VERSION : 0.1
   VAR_TEMP
      Pump_A : Struct
         Cond_01 : Bool;   // Condition 01
         Cond_02 : Bool;
         Cond_03 : Bool;   // Condition 03
      END_STRUCT;
      Pump_B : Struct
         Cond_01 : Bool;   // Condition 01
         Cond_02 : Bool;   // Condition 02
         Cond_03 : Bool;   // Condition 03
      END_STRUCT;
   END_VAR
BEGIN
   //****** Equipmens Activation*******
   //
   //IF "AlwaysFALSE" THEN
       //**************************************************************
       //Feed Water Pump A
       // Condition to CmdOn "On Command" 
       IF "P-104A_DB".Config.HMI.Enable_HMI_Controls = 1 THEN
           #Pump_A.Cond_01 := "T-104_DB".Equipments."P-104A".Enable AND ("T-104_DB".PmpSel."P-104AB" = 1 OR "T-104_DB".PmpSel."P-104AB" = 3);
           #Pump_A.Cond_02 := "T-104_DB".ExchangeCmds.Receive.ReqWater; //Route Open to sent to the Reactor
           "T-104_DB".Equipments."P-104A".CmdOn := #Pump_A.Cond_01 AND #Pump_A.Cond_02 AND NOT "T-104_DB".Cmds.Hold;
           IF "T-104_DB".Equipments."P-104A".CmdOn THEN
               "P-104A_DB".Stop_CMD := False;
               "P-104A_DB".Start_CMD := true;
               "P-104A_DB".ON := TRUE;
               "P-104A_DB".OFF := FALSE;
           ELSE
               "P-104A_DB".Stop_CMD := true;
               "P-104A_DB".Start_CMD := false;
               "P-104A_DB".ON := FALSE;
               "P-104A_DB".OFF := TRUE;
           END_IF;
       END_IF;
       //**************************************************************
       //Feed Water Pump B
       // Condition to CmdOn "On Command" 
       IF "P-104B_DB".Config.HMI.Enable_HMI_Controls = 1 THEN
           #Pump_B.Cond_01 := "T-104_DB".Equipments."P-104B".Enable AND ("T-104_DB".PmpSel."P-104AB" = 2 OR "T-104_DB".PmpSel."P-104AB" = 3);
           #Pump_B.Cond_02 := "T-104_DB".ExchangeCmds.Receive.ReqWater; //Route Open to sent to the Reactor
           "T-104_DB".Equipments."P-104B".CmdOn := #Pump_B.Cond_01 AND #Pump_B.Cond_02 AND NOT "T-104_DB".Cmds.Hold AND "AlwaysFALSE";
           IF "T-104_DB".Equipments."P-104B".CmdOn THEN
               "P-104B_DB".ON := TRUE;
               "P-104B_DB".OFF := FALSE;
           ELSE
               "P-104B_DB".ON := FALSE;
               "P-104B_DB".OFF := TRUE;
           END_IF;
       END_IF;
   //END_IF;
   "T-104_DB".ExchangeCmds.Send.PumpingOut := ("P-104A_DB".CF AND ("PT-104A_DB".SAI>0.2)) OR ("P-104B_DB".CF AND ("PT-104B_DB".SAI>0.2));
   "T-104_DB".ExchangeCmds.Send.PumpsOff := NOT "P-104A_DB".CF AND NOT "P-104B_DB".CF;//AND ("PT-104A_DB".SAI<0.2)) AND (NOT "P-104B_DB".CF AND ("PT-104B_DB".SAI<0.2));
   //*****************************************Tank Ready********************************************************************
   "T-104_DB".ExchangeCmds.Send.TankReady := "T-104_DB".Status.Step = 21 AND "T-104_DB".PmpSel."P-104AB" > 0;
END_FUNCTION

FUNCTION "T-104_SignalsOutExchange" : Void   // FC87, LAD
{ S7_Optimized_Access := 'TRUE' }
VERSION : 0.1
BEGIN

REGION Network 1: Started (Send)
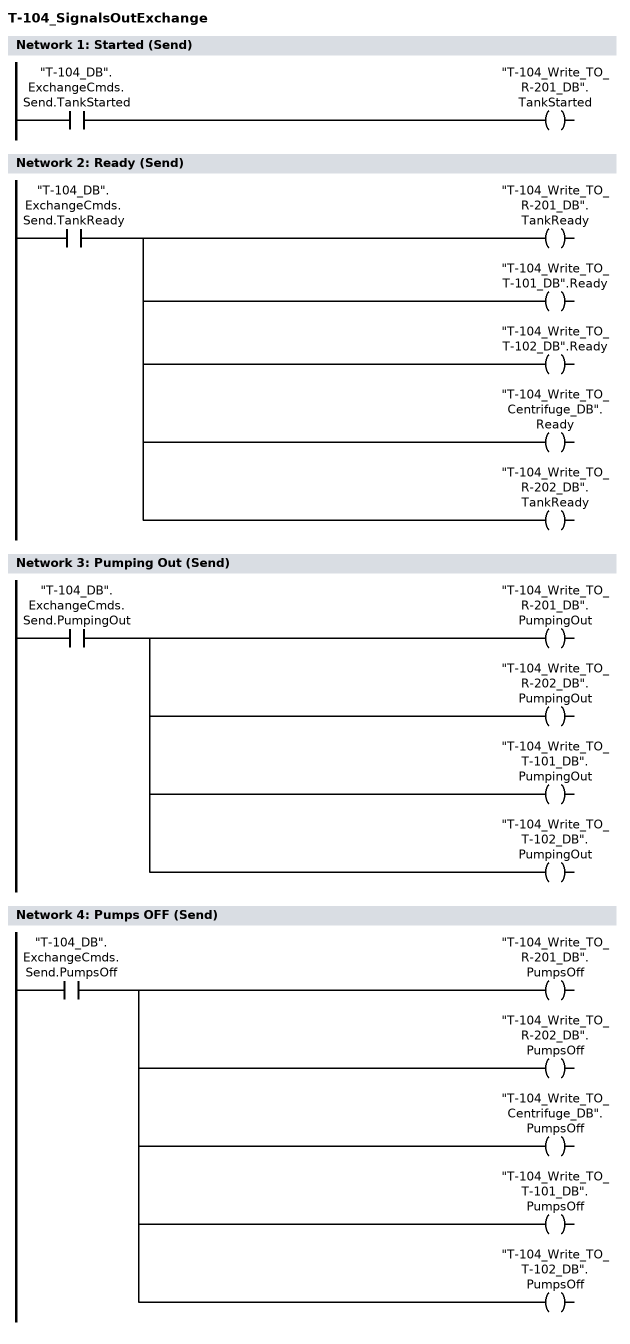
   RUNG wire#powerrail
      Contact( "T-104_DB".ExchangeCmds.Send.TankStarted )
      Coil( "T-104_Write_TO_R-201_DB".TankStarted )
   END_RUNG
   // the same network as SCL:
   "T-104_Write_TO_R-201_DB".TankStarted := "T-104_DB".ExchangeCmds.Send.TankStarted;
END_REGION

REGION Network 2: Ready (Send)
   RUNG wire#powerrail
      Contact( "T-104_DB".ExchangeCmds.Send.TankReady )
      wire#w1
      Coil( "T-104_Write_TO_R-201_DB".TankReady )
   END_RUNG
   RUNG wire#w1
      Coil( "T-104_Write_TO_T-101_DB".Ready )
   END_RUNG
   RUNG wire#w1
      Coil( "T-104_Write_TO_T-102_DB".Ready )
   END_RUNG
   RUNG wire#w1
      Coil( "T-104_Write_TO_Centrifuge_DB".Ready )
   END_RUNG
   RUNG wire#w1
      Coil( "T-104_Write_TO_R-202_DB".TankReady )
   END_RUNG
   // the same network as SCL:
   "T-104_Write_TO_R-201_DB".TankReady := "T-104_DB".ExchangeCmds.Send.TankReady;
   "T-104_Write_TO_T-101_DB".Ready := "T-104_DB".ExchangeCmds.Send.TankReady;
   "T-104_Write_TO_T-102_DB".Ready := "T-104_DB".ExchangeCmds.Send.TankReady;
   "T-104_Write_TO_Centrifuge_DB".Ready := "T-104_DB".ExchangeCmds.Send.TankReady;
   "T-104_Write_TO_R-202_DB".TankReady := "T-104_DB".ExchangeCmds.Send.TankReady;
END_REGION

REGION Network 3: Pumping Out (Send)
   RUNG wire#powerrail
      Contact( "T-104_DB".ExchangeCmds.Send.PumpingOut )
      wire#w1
      Coil( "T-104_Write_TO_R-201_DB".PumpingOut )
   END_RUNG
   RUNG wire#w1
      Coil( "T-104_Write_TO_R-202_DB".PumpingOut )
   END_RUNG
   RUNG wire#w1
      Coil( "T-104_Write_TO_T-101_DB".PumpingOut )
   END_RUNG
   RUNG wire#w1
      Coil( "T-104_Write_TO_T-102_DB".PumpingOut )
   END_RUNG
   // the same network as SCL:
   "T-104_Write_TO_R-201_DB".PumpingOut := "T-104_DB".ExchangeCmds.Send.PumpingOut;
   "T-104_Write_TO_R-202_DB".PumpingOut := "T-104_DB".ExchangeCmds.Send.PumpingOut;
   "T-104_Write_TO_T-101_DB".PumpingOut := "T-104_DB".ExchangeCmds.Send.PumpingOut;
   "T-104_Write_TO_T-102_DB".PumpingOut := "T-104_DB".ExchangeCmds.Send.PumpingOut;
END_REGION

REGION Network 4: Pumps OFF (Send)
   RUNG wire#powerrail
      Contact( "T-104_DB".ExchangeCmds.Send.PumpsOff )
      wire#w1
      Coil( "T-104_Write_TO_R-201_DB".PumpsOff )
   END_RUNG
   RUNG wire#w1
      Coil( "T-104_Write_TO_R-202_DB".PumpsOff )
   END_RUNG
   RUNG wire#w1
      Coil( "T-104_Write_TO_Centrifuge_DB".PumpsOff )
   END_RUNG
   RUNG wire#w1
      Coil( "T-104_Write_TO_T-101_DB".PumpsOff )
   END_RUNG
   RUNG wire#w1
      Coil( "T-104_Write_TO_T-102_DB".PumpsOff )
   END_RUNG
   // the same network as SCL:
   "T-104_Write_TO_R-201_DB".PumpsOff := "T-104_DB".ExchangeCmds.Send.PumpsOff;
   "T-104_Write_TO_R-202_DB".PumpsOff := "T-104_DB".ExchangeCmds.Send.PumpsOff;
   "T-104_Write_TO_Centrifuge_DB".PumpsOff := "T-104_DB".ExchangeCmds.Send.PumpsOff;
   "T-104_Write_TO_T-101_DB".PumpsOff := "T-104_DB".ExchangeCmds.Send.PumpsOff;
   "T-104_Write_TO_T-102_DB".PumpsOff := "T-104_DB".ExchangeCmds.Send.PumpsOff;
END_REGION
END_FUNCTION

FUNCTION "T-104_SEQ_FC" : Void   // FC88, LAD
{ S7_Optimized_Access := 'TRUE' }
VERSION : 0.1
   VAR_TEMP   // added for the SCL form of the ladder/FBD networks
      _w1 : Bool;
   END_VAR
BEGIN

REGION Network 2: Abort
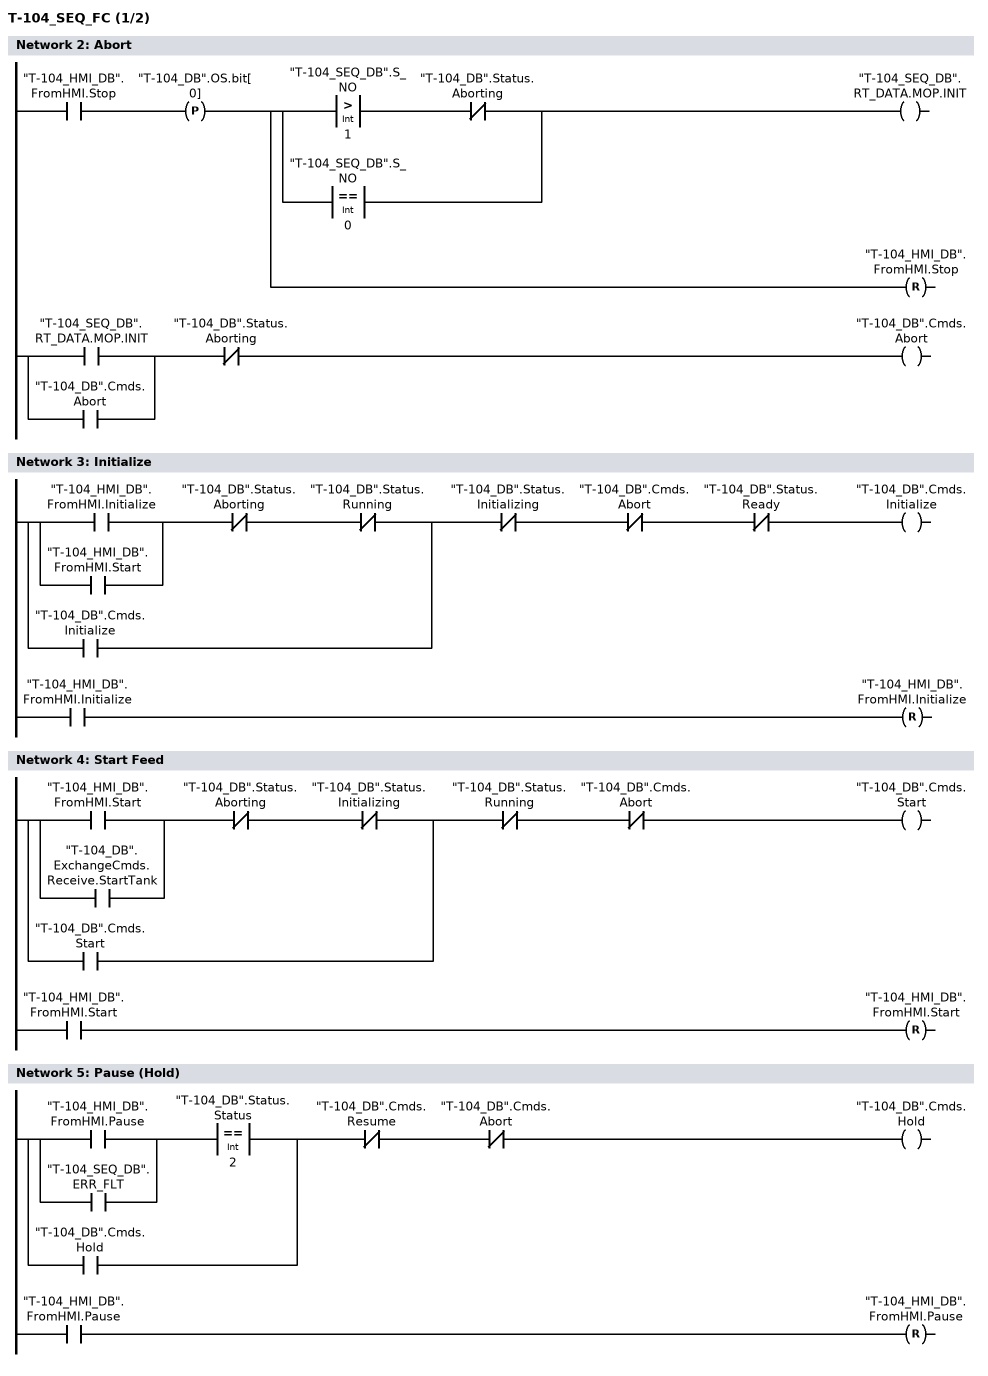
   RUNG wire#powerrail
      Contact( "T-104_HMI_DB".FromHMI.Stop )
      P_Trig( "T-104_DB".OS.bit[0] )
      wire#w1
      { S7_Templates := "SrcType := Int" } GT_Contact(in1 := "T-104_SEQ_DB".S_NO, in2 := 1)
      I_Contact( "T-104_DB".Status.Aborting )
      wire#w2
      Coil( "T-104_SEQ_DB".RT_DATA.MOP.INIT )
   END_RUNG
   RUNG wire#w1
      { S7_Templates := "SrcType := Int" } EQ_Contact(in1 := "T-104_SEQ_DB".S_NO, in2 := 0)
   END_RUNG wire#w2
   RUNG wire#w1
      R_Coil( "T-104_HMI_DB".FromHMI.Stop )
   END_RUNG
   RUNG wire#powerrail
      Contact( "T-104_SEQ_DB".RT_DATA.MOP.INIT )
      wire#w3
      I_Contact( "T-104_DB".Status.Aborting )
      Coil( "T-104_DB".Cmds.Abort )
   END_RUNG
   RUNG wire#powerrail
      Contact( "T-104_DB".Cmds.Abort )
   END_RUNG wire#w3
   // the same network as SCL:
   #_w1 := "T-104_HMI_DB".FromHMI.Stop AND NOT "T-104_DB".OS.bit[0];   // rising edge
   "T-104_DB".OS.bit[0] := "T-104_HMI_DB".FromHMI.Stop;
   "T-104_SEQ_DB".RT_DATA.MOP.INIT := #_w1 AND ((("T-104_SEQ_DB".S_NO > 1) AND NOT "T-104_DB".Status.Aborting) OR ("T-104_SEQ_DB".S_NO = 0));
   IF #_w1 THEN "T-104_HMI_DB".FromHMI.Stop := FALSE; END_IF;
   "T-104_DB".Cmds.Abort := ("T-104_SEQ_DB".RT_DATA.MOP.INIT OR "T-104_DB".Cmds.Abort) AND NOT "T-104_DB".Status.Aborting;
END_REGION

REGION Network 3: Initialize
   RUNG wire#powerrail
      Contact( "T-104_HMI_DB".FromHMI.Initialize )
      wire#w1
      I_Contact( "T-104_DB".Status.Aborting )
      I_Contact( "T-104_DB".Status.Running )
      wire#w2
      I_Contact( "T-104_DB".Status.Initializing )
      I_Contact( "T-104_DB".Cmds.Abort )
      I_Contact( "T-104_DB".Status.Ready )
      Coil( "T-104_DB".Cmds.Initialize )
   END_RUNG
   RUNG wire#powerrail
      Contact( "T-104_HMI_DB".FromHMI.Start )
   END_RUNG wire#w1
   RUNG wire#powerrail
      Contact( "T-104_DB".Cmds.Initialize )
   END_RUNG wire#w2
   RUNG wire#powerrail
      Contact( "T-104_HMI_DB".FromHMI.Initialize )
      R_Coil( "T-104_HMI_DB".FromHMI.Initialize )
   END_RUNG
   // the same network as SCL:
   "T-104_DB".Cmds.Initialize := ((("T-104_HMI_DB".FromHMI.Initialize OR "T-104_HMI_DB".FromHMI.Start) AND NOT "T-104_DB".Status.Aborting AND NOT "T-104_DB".Status.Running) OR "T-104_DB".Cmds.Initialize) AND NOT "T-104_DB".Status.Initializing AND NOT "T-104_DB".Cmds.Abort AND NOT "T-104_DB".Status.Ready;
   IF "T-104_HMI_DB".FromHMI.Initialize THEN "T-104_HMI_DB".FromHMI.Initialize := FALSE; END_IF;
END_REGION

REGION Network 4: Start Feed
   RUNG wire#powerrail
      Contact( "T-104_HMI_DB".FromHMI.Start )
      wire#w1
      I_Contact( "T-104_DB".Status.Aborting )
      I_Contact( "T-104_DB".Status.Initializing )
      wire#w2
      I_Contact( "T-104_DB".Status.Running )
      I_Contact( "T-104_DB".Cmds.Abort )
      Coil( "T-104_DB".Cmds.Start )
   END_RUNG
   RUNG wire#powerrail
      Contact( "T-104_DB".ExchangeCmds.Receive.StartTank )
   END_RUNG wire#w1
   RUNG wire#powerrail
      Contact( "T-104_DB".Cmds.Start )
   END_RUNG wire#w2
   RUNG wire#powerrail
      Contact( "T-104_HMI_DB".FromHMI.Start )
      R_Coil( "T-104_HMI_DB".FromHMI.Start )
   END_RUNG
   // the same network as SCL:
   "T-104_DB".Cmds.Start := ((("T-104_HMI_DB".FromHMI.Start OR "T-104_DB".ExchangeCmds.Receive.StartTank) AND NOT "T-104_DB".Status.Aborting AND NOT "T-104_DB".Status.Initializing) OR "T-104_DB".Cmds.Start) AND NOT "T-104_DB".Status.Running AND NOT "T-104_DB".Cmds.Abort;
   IF "T-104_HMI_DB".FromHMI.Start THEN "T-104_HMI_DB".FromHMI.Start := FALSE; END_IF;
END_REGION

REGION Network 5: Pause (Hold)
   RUNG wire#powerrail
      Contact( "T-104_HMI_DB".FromHMI.Pause )
      wire#w1
      { S7_Templates := "SrcType := Int" } EQ_Contact(in1 := "T-104_DB".Status.Status, in2 := 2)
      wire#w2
      I_Contact( "T-104_DB".Cmds.Resume )
      I_Contact( "T-104_DB".Cmds.Abort )
      Coil( "T-104_DB".Cmds.Hold )
   END_RUNG
   RUNG wire#powerrail
      Contact( "T-104_SEQ_DB".ERR_FLT )
   END_RUNG wire#w1
   RUNG wire#powerrail
      Contact( "T-104_DB".Cmds.Hold )
   END_RUNG wire#w2
   RUNG wire#powerrail
      Contact( "T-104_HMI_DB".FromHMI.Pause )
      R_Coil( "T-104_HMI_DB".FromHMI.Pause )
   END_RUNG
   // the same network as SCL:
   "T-104_DB".Cmds.Hold := ((("T-104_HMI_DB".FromHMI.Pause OR "T-104_SEQ_DB".ERR_FLT) AND ("T-104_DB".Status.Status = 2)) OR "T-104_DB".Cmds.Hold) AND NOT "T-104_DB".Cmds.Resume AND NOT "T-104_DB".Cmds.Abort;
   IF "T-104_HMI_DB".FromHMI.Pause THEN "T-104_HMI_DB".FromHMI.Pause := FALSE; END_IF;
END_REGION

REGION Network 6: Restart From Pause (Hold)
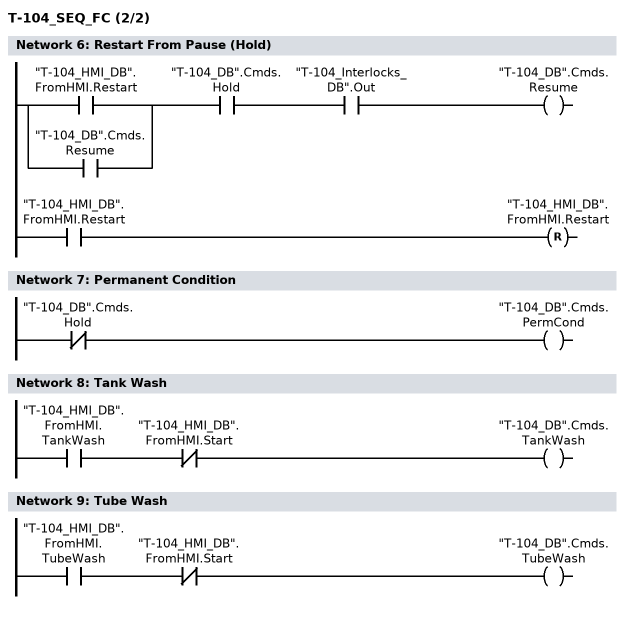
   RUNG wire#powerrail
      Contact( "T-104_HMI_DB".FromHMI.Restart )
      wire#w1
      Contact( "T-104_DB".Cmds.Hold )
      Contact( "T-104_Interlocks_DB".Out )
      Coil( "T-104_DB".Cmds.Resume )
   END_RUNG
   RUNG wire#powerrail
      Contact( "T-104_DB".Cmds.Resume )
   END_RUNG wire#w1
   RUNG wire#powerrail
      Contact( "T-104_HMI_DB".FromHMI.Restart )
      R_Coil( "T-104_HMI_DB".FromHMI.Restart )
   END_RUNG
   // the same network as SCL:
   "T-104_DB".Cmds.Resume := ("T-104_HMI_DB".FromHMI.Restart OR "T-104_DB".Cmds.Resume) AND "T-104_DB".Cmds.Hold AND "T-104_Interlocks_DB".Out;
   IF "T-104_HMI_DB".FromHMI.Restart THEN "T-104_HMI_DB".FromHMI.Restart := FALSE; END_IF;
END_REGION

REGION Network 7: Permanent Condition
   RUNG wire#powerrail
      I_Contact( "T-104_DB".Cmds.Hold )
      Coil( "T-104_DB".Cmds.PermCond )
   END_RUNG
   // the same network as SCL:
   "T-104_DB".Cmds.PermCond := NOT "T-104_DB".Cmds.Hold;
END_REGION

REGION Network 8: Tank Wash
   RUNG wire#powerrail
      Contact( "T-104_HMI_DB".FromHMI.TankWash )
      I_Contact( "T-104_HMI_DB".FromHMI.Start )
      Coil( "T-104_DB".Cmds.TankWash )
   END_RUNG
   // the same network as SCL:
   "T-104_DB".Cmds.TankWash := "T-104_HMI_DB".FromHMI.TankWash AND NOT "T-104_HMI_DB".FromHMI.Start;
END_REGION

REGION Network 9: Tube Wash
   RUNG wire#powerrail
      Contact( "T-104_HMI_DB".FromHMI.TubeWash )
      I_Contact( "T-104_HMI_DB".FromHMI.Start )
      Coil( "T-104_DB".Cmds.TubeWash )
   END_RUNG
   // the same network as SCL:
   "T-104_DB".Cmds.TubeWash := "T-104_HMI_DB".FromHMI.TubeWash AND NOT "T-104_HMI_DB".FromHMI.Start;
END_REGION

REGION Network 10 (SCL): Sequence Status
   IF "T-104_SEQ_DB".S_NO= 1 THEN
       "T-104_DB".Status.Status := 1; //Idle
   ELSIF "T-104_SEQ_DB".S_NO > 1 AND "T-104_SEQ_DB".S_NO < 150 AND NOT "T-104_SEQ_DB".ERR_FLT AND NOT "T-104_DB".Cmds.Hold THEN
       "T-104_DB".Status.Status := 2; //Running
   ELSIF "T-104_SEQ_DB".S_NO >= 151 AND "T-104_SEQ_DB".S_NO <= 160 AND NOT "T-104_SEQ_DB".ERR_FLT THEN
       "T-104_DB".Status.Status := 3; // Stopping
   ELSIF  "T-104_SEQ_DB".ERR_FLT AND  ("T-104_SEQ_DB".S_NO > 1 AND "T-104_SEQ_DB".S_NO < 150) THEN
       "T-104_DB".Status.Status := 4; // Held
   ELSIF  "T-104_SEQ_DB".ERR_FLT AND  ("T-104_SEQ_DB".S_NO > 1 AND "T-104_SEQ_DB".S_NO < 150) AND "T-104_Aux_DB"."Bool".TOff  THEN
       "T-104_DB".Status.Status := 5; // Holding
   ELSE
       "T-104_DB".Status.Status := 6; // Unknown
   END_IF;

   "T-104_DB".Status.Running := ("T-104_SEQ_DB".S_NO > 3 AND "T-104_SEQ_DB".S_NO <= 150);
   "T-104_DB".Status.Initializing := ("T-104_SEQ_DB".S_NO >= 141 AND "T-104_SEQ_DB".S_NO <= 150);

   //Enable/Disable HMI Start/Stop Button
   "T-104_HMI_DB".ToHMI.EnStopButton := ("T-104_DB".Status.Status > 1) OR "T-104_DB".Status.Step = 0; //Enable HMI Stop Button
   "T-104_HMI_DB".ToHMI.EnStartButton := "T-104_DB".Status.Status = 1; //Idle
   "T-104_HMI_DB".ToHMI.EnPauseButton := "T-104_DB".Status.Status = 2; //Enable Pause Button
   "T-104_HMI_DB".ToHMI.EnRestartButton :=  "T-104_DB".Status.Status = 4; //Enable Restart Button

   //****Interlock Activated
   "T-104_HMI_DB".ToHMI.InterlockActivated := "T-104_Interlocks_DB".Out;
END_REGION

REGION Network 11 (SCL): Sequence Step
   "T-104_DB".Status.Step := "T-104_SEQ_DB".S_NO;
END_REGION

REGION Network 12 (SCL): Sequence state (Procedure running)
   IF "T-104_SEQ_DB".S_NO = 3 OR "T-104_SEQ_DB".S_NO = 4 THEN
       "T-104_DB".Status.State := 1; //Ready
   ELSIF "T-104_SEQ_DB".S_NO >= 21 AND "T-104_SEQ_DB".S_NO <= 60 THEN
       "T-104_DB".Status.State := 2; //Mixing 
   ELSIF "T-104_SEQ_DB".S_NO >= 61 AND "T-104_SEQ_DB".S_NO <= 80 THEN
       "T-104_DB".Status.State := 3; //Pouring
   ELSIF "T-104_SEQ_DB".S_NO >= 141 AND "T-104_SEQ_DB".S_NO <= 150 THEN
       "T-104_DB".Status.State := 4; //Initializing
   ELSIF "T-104_SEQ_DB".S_NO >= 151 AND "T-104_SEQ_DB".S_NO <= 160 THEN
       "T-104_DB".Status.State := 5; //Aborting
   ELSE
       "T-104_DB".Status.State := 0;
   END_IF;
END_REGION

REGION Network 13: Sequence State
END_REGION
END_FUNCTION

// folder: State MACHINE/1)Tanks/Tank T-104 (Water System)/T-104 <---> Centrifuge

FUNCTION "T-104_Signals_FROM_Centrifuge" : Void   // FC71, LAD
{ S7_Optimized_Access := 'TRUE' }
VERSION : 0.1
BEGIN

REGION Network 1: Start Sequence
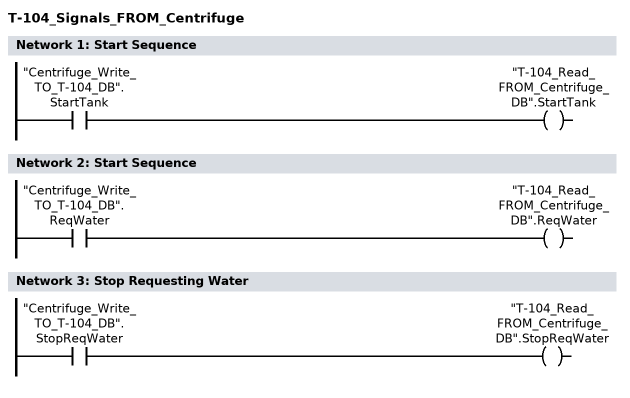
   RUNG wire#powerrail
      Contact( "Centrifuge_Write_TO_T-104_DB".StartTank )
      Coil( "T-104_Read_FROM_Centrifuge_DB".StartTank )
   END_RUNG
   // the same network as SCL:
   "T-104_Read_FROM_Centrifuge_DB".StartTank := "Centrifuge_Write_TO_T-104_DB".StartTank;
END_REGION

REGION Network 2: Start Sequence
   RUNG wire#powerrail
      Contact( "Centrifuge_Write_TO_T-104_DB".ReqWater )
      Coil( "T-104_Read_FROM_Centrifuge_DB".ReqWater )
   END_RUNG
   // the same network as SCL:
   "T-104_Read_FROM_Centrifuge_DB".ReqWater := "Centrifuge_Write_TO_T-104_DB".ReqWater;
END_REGION

REGION Network 3: Stop Requesting Water
   RUNG wire#powerrail
      Contact( "Centrifuge_Write_TO_T-104_DB".StopReqWater )
      Coil( "T-104_Read_FROM_Centrifuge_DB".StopReqWater )
   END_RUNG
   // the same network as SCL:
   "T-104_Read_FROM_Centrifuge_DB".StopReqWater := "Centrifuge_Write_TO_T-104_DB".StopReqWater;
END_REGION
END_FUNCTION

// folder: State MACHINE/1)Tanks/Tank T-104 (Water System)/T-104 <---> R-201

FUNCTION "T-104_Signals_FROM_R-201" : Void   // FC50, LAD
{ S7_Optimized_Access := 'TRUE' }
VERSION : 0.1
BEGIN

REGION Network 1: Start Sequence
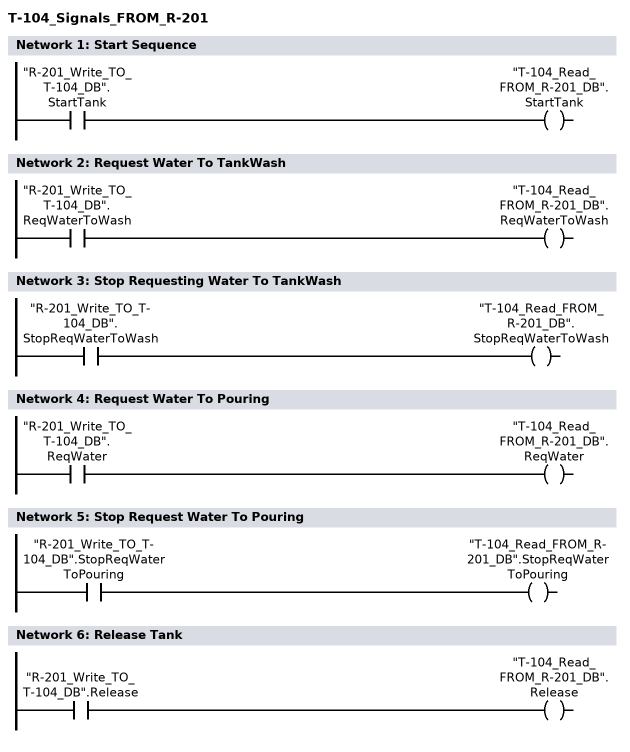
   RUNG wire#powerrail
      Contact( "R-201_Write_TO_T-104_DB".StartTank )
      Coil( "T-104_Read_FROM_R-201_DB".StartTank )
   END_RUNG
   // the same network as SCL:
   "T-104_Read_FROM_R-201_DB".StartTank := "R-201_Write_TO_T-104_DB".StartTank;
END_REGION

REGION Network 2: Request Water To TankWash
   RUNG wire#powerrail
      Contact( "R-201_Write_TO_T-104_DB".ReqWaterToWash )
      Coil( "T-104_Read_FROM_R-201_DB".ReqWaterToWash )
   END_RUNG
   // the same network as SCL:
   "T-104_Read_FROM_R-201_DB".ReqWaterToWash := "R-201_Write_TO_T-104_DB".ReqWaterToWash;
END_REGION

REGION Network 3: Stop Requesting Water To TankWash
   RUNG wire#powerrail
      Contact( "R-201_Write_TO_T-104_DB".StopReqWaterToWash )
      Coil( "T-104_Read_FROM_R-201_DB".StopReqWaterToWash )
   END_RUNG
   // the same network as SCL:
   "T-104_Read_FROM_R-201_DB".StopReqWaterToWash := "R-201_Write_TO_T-104_DB".StopReqWaterToWash;
END_REGION

REGION Network 4: Request Water To Pouring
   RUNG wire#powerrail
      Contact( "R-201_Write_TO_T-104_DB".ReqWater )
      Coil( "T-104_Read_FROM_R-201_DB".ReqWater )
   END_RUNG
   // the same network as SCL:
   "T-104_Read_FROM_R-201_DB".ReqWater := "R-201_Write_TO_T-104_DB".ReqWater;
END_REGION

REGION Network 5: Stop Request Water To Pouring
   RUNG wire#powerrail
      Contact( "R-201_Write_TO_T-104_DB".StopReqWaterToPouring )
      Coil( "T-104_Read_FROM_R-201_DB".StopReqWaterToPouring )
   END_RUNG
   // the same network as SCL:
   "T-104_Read_FROM_R-201_DB".StopReqWaterToPouring := "R-201_Write_TO_T-104_DB".StopReqWaterToPouring;
END_REGION

REGION Network 6: Release Tank
   RUNG wire#powerrail
      Contact( "R-201_Write_TO_T-104_DB".Release )
      Coil( "T-104_Read_FROM_R-201_DB".Release )
   END_RUNG
   // the same network as SCL:
   "T-104_Read_FROM_R-201_DB".Release := "R-201_Write_TO_T-104_DB".Release;
END_REGION
END_FUNCTION

// folder: State MACHINE/1)Tanks/Tank T-104 (Water System)/T-104 <---> R-202

FUNCTION "T-104_Signals_FROM_R-202" : Void   // FC72, LAD
{ S7_Optimized_Access := 'TRUE' }
VERSION : 0.1
BEGIN

REGION Network 1: Start Sequence
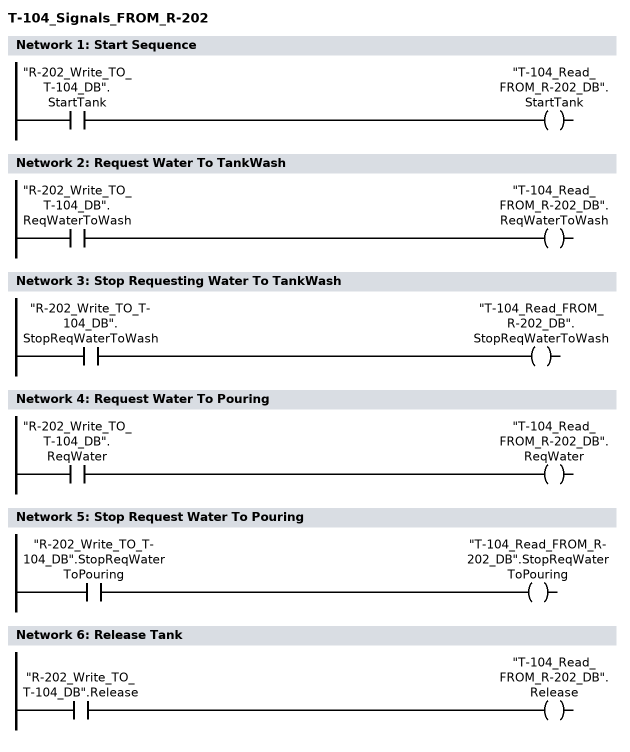
   RUNG wire#powerrail
      Contact( "R-202_Write_TO_T-104_DB".StartTank )
      Coil( "T-104_Read_FROM_R-202_DB".StartTank )
   END_RUNG
   // the same network as SCL:
   "T-104_Read_FROM_R-202_DB".StartTank := "R-202_Write_TO_T-104_DB".StartTank;
END_REGION

REGION Network 2: Request Water To TankWash
   RUNG wire#powerrail
      Contact( "R-202_Write_TO_T-104_DB".ReqWaterToWash )
      Coil( "T-104_Read_FROM_R-202_DB".ReqWaterToWash )
   END_RUNG
   // the same network as SCL:
   "T-104_Read_FROM_R-202_DB".ReqWaterToWash := "R-202_Write_TO_T-104_DB".ReqWaterToWash;
END_REGION

REGION Network 3: Stop Requesting Water To TankWash
   RUNG wire#powerrail
      Contact( "R-202_Write_TO_T-104_DB".StopReqWaterToWash )
      Coil( "T-104_Read_FROM_R-202_DB".StopReqWaterToWash )
   END_RUNG
   // the same network as SCL:
   "T-104_Read_FROM_R-202_DB".StopReqWaterToWash := "R-202_Write_TO_T-104_DB".StopReqWaterToWash;
END_REGION

REGION Network 4: Request Water To Pouring
   RUNG wire#powerrail
      Contact( "R-202_Write_TO_T-104_DB".ReqWater )
      Coil( "T-104_Read_FROM_R-202_DB".ReqWater )
   END_RUNG
   // the same network as SCL:
   "T-104_Read_FROM_R-202_DB".ReqWater := "R-202_Write_TO_T-104_DB".ReqWater;
END_REGION

REGION Network 5: Stop Request Water To Pouring
   RUNG wire#powerrail
      Contact( "R-202_Write_TO_T-104_DB".StopReqWaterToPouring )
      Coil( "T-104_Read_FROM_R-202_DB".StopReqWaterToPouring )
   END_RUNG
   // the same network as SCL:
   "T-104_Read_FROM_R-202_DB".StopReqWaterToPouring := "R-202_Write_TO_T-104_DB".StopReqWaterToPouring;
END_REGION

REGION Network 6: Release Tank
   RUNG wire#powerrail
      Contact( "R-202_Write_TO_T-104_DB".Release )
      Coil( "T-104_Read_FROM_R-202_DB".Release )
   END_RUNG
   // the same network as SCL:
   "T-104_Read_FROM_R-202_DB".Release := "R-202_Write_TO_T-104_DB".Release;
END_REGION
END_FUNCTION

// folder: State MACHINE/1)Tanks/Tank T-104 (Water System)/T-104 <---> T-101

FUNCTION "T-104_Signals_FROM_T-101" : Void   // FC74, LAD
{ S7_Optimized_Access := 'TRUE' }
VERSION : 0.1
BEGIN

REGION Network 1: Start Sequence
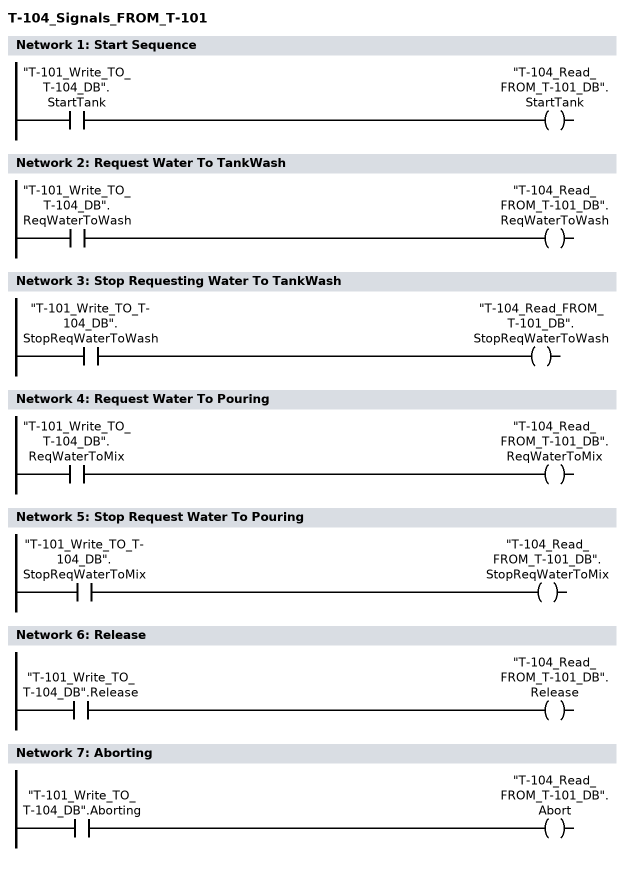
   RUNG wire#powerrail
      Contact( "T-101_Write_TO_T-104_DB".StartTank )
      Coil( "T-104_Read_FROM_T-101_DB".StartTank )
   END_RUNG
   // the same network as SCL:
   "T-104_Read_FROM_T-101_DB".StartTank := "T-101_Write_TO_T-104_DB".StartTank;
END_REGION

REGION Network 2: Request Water To TankWash
   RUNG wire#powerrail
      Contact( "T-101_Write_TO_T-104_DB".ReqWaterToWash )
      Coil( "T-104_Read_FROM_T-101_DB".ReqWaterToWash )
   END_RUNG
   // the same network as SCL:
   "T-104_Read_FROM_T-101_DB".ReqWaterToWash := "T-101_Write_TO_T-104_DB".ReqWaterToWash;
END_REGION

REGION Network 3: Stop Requesting Water To TankWash
   RUNG wire#powerrail
      Contact( "T-101_Write_TO_T-104_DB".StopReqWaterToWash )
      Coil( "T-104_Read_FROM_T-101_DB".StopReqWaterToWash )
   END_RUNG
   // the same network as SCL:
   "T-104_Read_FROM_T-101_DB".StopReqWaterToWash := "T-101_Write_TO_T-104_DB".StopReqWaterToWash;
END_REGION

REGION Network 4: Request Water To Pouring
   RUNG wire#powerrail
      Contact( "T-101_Write_TO_T-104_DB".ReqWaterToMix )
      Coil( "T-104_Read_FROM_T-101_DB".ReqWaterToMix )
   END_RUNG
   // the same network as SCL:
   "T-104_Read_FROM_T-101_DB".ReqWaterToMix := "T-101_Write_TO_T-104_DB".ReqWaterToMix;
END_REGION

REGION Network 5: Stop Request Water To Pouring
   RUNG wire#powerrail
      Contact( "T-101_Write_TO_T-104_DB".StopReqWaterToMix )
      Coil( "T-104_Read_FROM_T-101_DB".StopReqWaterToMix )
   END_RUNG
   // the same network as SCL:
   "T-104_Read_FROM_T-101_DB".StopReqWaterToMix := "T-101_Write_TO_T-104_DB".StopReqWaterToMix;
END_REGION

REGION Network 6: Release
   RUNG wire#powerrail
      Contact( "T-101_Write_TO_T-104_DB".Release )
      Coil( "T-104_Read_FROM_T-101_DB".Release )
   END_RUNG
   // the same network as SCL:
   "T-104_Read_FROM_T-101_DB".Release := "T-101_Write_TO_T-104_DB".Release;
END_REGION

REGION Network 7: Aborting
   RUNG wire#powerrail
      Contact( "T-101_Write_TO_T-104_DB".Aborting )
      Coil( "T-104_Read_FROM_T-101_DB".Abort )
   END_RUNG
   // the same network as SCL:
   "T-104_Read_FROM_T-101_DB".Abort := "T-101_Write_TO_T-104_DB".Aborting;
END_REGION
END_FUNCTION

// folder: State MACHINE/1)Tanks/Tank T-104 (Water System)/T-104 <---> T-102

FUNCTION "T-104_Signals_FROM_T-102" : Void   // FC73, LAD
{ S7_Optimized_Access := 'TRUE' }
VERSION : 0.1
BEGIN

REGION Network 1: Start Sequence
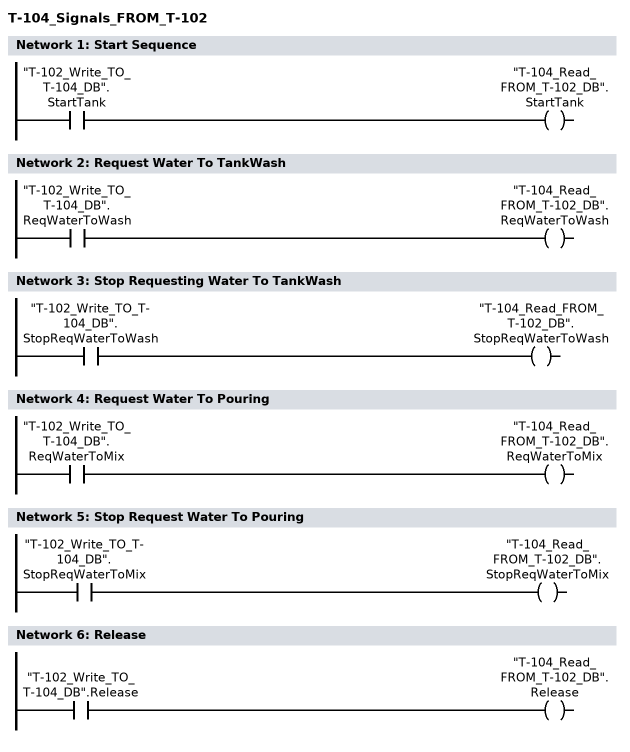
   RUNG wire#powerrail
      Contact( "T-102_Write_TO_T-104_DB".StartTank )
      Coil( "T-104_Read_FROM_T-102_DB".StartTank )
   END_RUNG
   // the same network as SCL:
   "T-104_Read_FROM_T-102_DB".StartTank := "T-102_Write_TO_T-104_DB".StartTank;
END_REGION

REGION Network 2: Request Water To TankWash
   RUNG wire#powerrail
      Contact( "T-102_Write_TO_T-104_DB".ReqWaterToWash )
      Coil( "T-104_Read_FROM_T-102_DB".ReqWaterToWash )
   END_RUNG
   // the same network as SCL:
   "T-104_Read_FROM_T-102_DB".ReqWaterToWash := "T-102_Write_TO_T-104_DB".ReqWaterToWash;
END_REGION

REGION Network 3: Stop Requesting Water To TankWash
   RUNG wire#powerrail
      Contact( "T-102_Write_TO_T-104_DB".StopReqWaterToWash )
      Coil( "T-104_Read_FROM_T-102_DB".StopReqWaterToWash )
   END_RUNG
   // the same network as SCL:
   "T-104_Read_FROM_T-102_DB".StopReqWaterToWash := "T-102_Write_TO_T-104_DB".StopReqWaterToWash;
END_REGION

REGION Network 4: Request Water To Pouring
   RUNG wire#powerrail
      Contact( "T-102_Write_TO_T-104_DB".ReqWaterToMix )
      Coil( "T-104_Read_FROM_T-102_DB".ReqWaterToMix )
   END_RUNG
   // the same network as SCL:
   "T-104_Read_FROM_T-102_DB".ReqWaterToMix := "T-102_Write_TO_T-104_DB".ReqWaterToMix;
END_REGION

REGION Network 5: Stop Request Water To Pouring
   RUNG wire#powerrail
      Contact( "T-102_Write_TO_T-104_DB".StopReqWaterToMix )
      Coil( "T-104_Read_FROM_T-102_DB".StopReqWaterToMix )
   END_RUNG
   // the same network as SCL:
   "T-104_Read_FROM_T-102_DB".StopReqWaterToMix := "T-102_Write_TO_T-104_DB".StopReqWaterToMix;
END_REGION

REGION Network 6: Release
   RUNG wire#powerrail
      Contact( "T-102_Write_TO_T-104_DB".Release )
      Coil( "T-104_Read_FROM_T-102_DB".Release )
   END_RUNG
   // the same network as SCL:
   "T-104_Read_FROM_T-102_DB".Release := "T-102_Write_TO_T-104_DB".Release;
END_REGION
END_FUNCTION

// folder: State MACHINE/2)Reactors/Reactor R-201

FUNCTION_BLOCK "R-201_SEQ"   // FB32, GRAPH_PLUS
{ S7_Optimized_Access := 'TRUE' }
VERSION : 0.1
   VAR_INPUT
      OFF_SQ : Bool := false;   // Turn sequence off
      INIT_SQ : Bool := false;   // Set sequence to initial state
      ACK_EF : Bool := false;   // Acknowledge all errors and faults
   END_VAR
   VAR_OUTPUT
      S_NO : Int := 0;   // Step number
      S_MORE : Bool := false;   // More steps are available and can be shown in S_NO
      S_ACTIVE : Bool := false;   // Step indicated in S_NO is active
      ERR_FLT : Bool := false;   // Interlock or supervision group error
      AUTO_ON : Bool := false;   // Automatic mode is active
   END_VAR
   VAR
      Reactor : Struct   // Reactor Ctrl
         IDLE : Bool;
         INITIALIZATION : Bool;   // Sequence initialization
         START : Bool;
         DONE_REACTING : Bool;
         COMPLETE : Bool;   // Reactor Complete Read only
         PARA : Bool;   // PARA load Batch side button
         ABORTING : Bool;   // Sequence about
         WAIT : Bool;   // Wating for Permissive read only
      END_STRUCT;
      "Aux Reactor" : Struct
         INITIALIZATION : Bool;
         START : Bool;
         DONE : Bool;
         COMPLETE : Bool;
         PARA : Bool;
         "SELECT_R-201" : Bool;
         "SELECT_R-202" : Bool;
         "SELECT_R-201/R-202" : Bool;
         "SELECT_R-201_T-103" : Bool;
         "SELECT_R-202_T-103" : Bool;
         ABORT : Bool;
         WAIT : Bool;
         LV : Bool;
         FLOW : Bool;
         MIX : Bool;
         "Pre-MIX" : Bool;
         REACTOR : Bool;
         WASH : Bool;
         TUBE : Bool;
         "SEQ_R-201" : Bool;
         "SEQ_R-202" : Bool;
         "SEQ_ R-201 & R-202" : Bool;
         "SEQ_T-103_R-201" : Bool;
         "SEQ_T-103_R-202" : Bool;
         BatchVolume : Real;
         Batchsize : Real;
         batchFlow : Real := 1.0;
         "batchFlow_T-102" : Real;
         BatchPH : Real := 7.0;
         "T-101" : Real;
         BatchTemp : Real := 80.0;
         PM : Bool;
         "TIME" : Struct
            "PRE-MIX" : Time;
            PH_DELAY : Time;
            REACTOR : Time;
            WATCH : Time;
            TUBE : Time;
            CountDown : Struct
               "PRE-MIX" : Time;
               PH_DELAY : Time;
               REACTOR : Time;
               WATCH : Time;
               TUBE : Time;
            END_STRUCT;
         END_STRUCT;
         "TIMER" : Struct
            "PRE-MIX" : IEC_TIMER;
            MIX : IEC_TIMER;
            PH_DELAY : IEC_TIMER;
            REACTOR : IEC_TIMER;
            WASH : IEC_TIMER;
            TUBE : IEC_TIMER;
         END_STRUCT;
      END_STRUCT;
      TEMP : Struct
         TANKS_BATCH : Real;
         "EMPTY_LV_0%" : Real;
         "MIN_LV_20%" : Real;
         "MAX_LV_80%" : Real;
         "BELOW_32%" : Real;
         "Greater_8%" : Real;
         "PRE-ADD" : Real;
         X_SOL_SIZE : Real;
         Y_SOL_SIZE : Real;
         PH_MIN : Real;
         PH_MAX : Real;
         OFFSEt : Struct
            MAX : Real;
            MIN : Real;
         END_STRUCT;
      END_STRUCT;
      COOLING : Struct   // Reactor Ctrl
         IDLE : Bool;
      END_STRUCT;
      HMI_INFO : Array[0..16] of UInt;
      IF_PAR : G7_IfParPlus_V6;
      RT_DATA : G7_RTDataPlus_V6;   // Internal data area
      Abort : G7_TransitionPlus_V6;   // Transition structure
      InitializeR : G7_TransitionPlus_V6;   // Transition structure
      "Fill/Pouring" : G7_TransitionPlus_V6;   // Transition structure
      Re : G7_TransitionPlus_V6;   // Transition structure
      "Fill/Pour" : G7_TransitionPlus_V6;   // Transition structure
      WashT : G7_TransitionPlus_V6;   // Transition structure
      WashTub : G7_TransitionPlus_V6;   // Transition structure
      Std : G7_TransitionPlus_V6;   // Transition structure
      StT : G7_TransitionPlus_V6;   // Transition structure
      WatFll : G7_TransitionPlus_V6;   // Transition structure
      StRW : G7_TransitionPlus_V6;   // Transition structure
      RelT : G7_TransitionPlus_V6;   // Transition structure
      PMix : G7_TransitionPlus_V6;   // Transition structure
      OpR : G7_TransitionPlus_V6;   // Transition structure
      TOT_Done : G7_TransitionPlus_V6;   // Transition structure
      PmpOFF : G7_TransitionPlus_V6;   // Transition structure
      IdleTank : G7_TransitionPlus_V6;   // Transition structure
      TS : G7_TransitionPlus_V6;   // Transition structure
      pHCtl : G7_TransitionPlus_V6;   // Transition structure
      pHCtl2 : G7_TransitionPlus_V6;   // Transition structure
      PmpOFF2 : G7_TransitionPlus_V6;   // Transition structure
      T102_Idle : G7_TransitionPlus_V6;   // Transition structure
      PourD : G7_TransitionPlus_V6;   // Transition structure